(* Logix 5000 project; controller MV vendor 1 type 14 code 217 rev 31.11; software revision 31.00; part 45 of 53 *)
(* tags used below, declared in another part *)
   Always_Off : BOOL;
   CWD : CHECKWORD_FLAGS;
   Enable_TimeString : BOOL;
   MV22_TP_Capture_Volume_Timer : TIMER;
   MV_BM01_AV01 : PlantItem;   // BM01_AV01
   MV_BM01_AV01_CIP : BOOL;
   MV_BM01_AV01_MV21 : BOOL;
   MV_DAL01_AV01_MV21 : BOOL;
   MV_Enable_MV21_NewPressureControl : BOOL;
   MV_Enable_MV22_NewPressureControl : BOOL;
   MV_GasAvailable : BOOL;
   MV_MV21_AV01 : PlantItem;   // MV21_AV01
   MV_MV21_CIP : BOOL;
   MV_MV21_CO2 : BOOL;
   MV_MV21_CO2_ON_PreStorage : BOOL;
   MV_MV21_CO2_ON_Storage : BOOL;
   MV_MV21_ControlOpenVent : BOOL;
   MV_MV21_Filling_Pulse : BOOL;
   MV_MV21_Filling_PulseLevel : REAL;
   MV_MV21_LTX07_TrueLevel : REAL;
   MV_MV21_ProxiesOK : BOOL;
   MV_MV21_PTX01_AI : PlantItem;   // MV21_PTX01
   MV_MV21_TP_CaskDepressure : BOOL;
   MV_MV21_TP_CaskEmptying : BOOL;
   MV_MV21_TP_CaskFilling : BOOL;
   MV_MV21_TP_CaskPrePressure : BOOL;
   MV_MV21_TP_CaskReadyToFill : BOOL;
   MV_MV21_TP_CaskStorage : BOOL;
   MV_MV21_TP_CO2_Debounce_Timer : TIMER;
   MV_MV21_TP_CO2_Debounce_Timer_1 : TIMER;
   MV_MV21_TP_CO2_HSL_Pressure : REAL;
   MV_MV21_TP_CO2_HSL_Storage : REAL;
   MV_MV21_TP_CO2_HSL_Timer : TIMER;
   MV_MV21_TP_CO2_LSL_pressure_1 : REAL;
   MV_MV21_TP_CO2_LSL_storage : REAL;
   MV_MV21_TP_CO2_LSL_Timer : TIMER;
   MV_MV21_TP_Command : DINT;
   MV_MV21_TP_DAL_Chase_Cask : BOOL;
   MV_MV21_TP_DAL_Chase_KB : BOOL;
   MV_MV21_TP_DAL_Chase_Time : TIMER;
   MV_MV21_TP_Error_String : STRING;
   MV_MV21_TP_Faulted : BOOL;
   MV_MV21_TP_Fill_Pulse_OFF_Timer : TIMER;
   MV_MV21_TP_Fill_Pulse_ON_Timer : TIMER;
   MV_MV21_TP_Held : BOOL;
   MV_MV21_TP_Idle : BOOL;
   MV_MV21_TP_Initial_DAL_Chase_Cask : BOOL;
   MV_MV21_TP_Initial_DAL_Chase_KB : BOOL;
   MV_MV21_TP_KBEmptying : BOOL;
   MV_MV21_TP_KBFilling : BOOL;
   MV_MV21_TP_KBFillingBuildPressure : BOOL;
   MV_MV21_TP_KBPreEmptyPressure : BOOL;
   MV_MV21_TP_KBPrePressurise : BOOL;
   MV_MV21_TP_KBStorage : BOOL;
   MV_MV21_TP_LowerLimit : REAL;
   MV_MV21_TP_NotIdle : BOOL;
   MV_MV21_TP_Prompt : DINT;
   MV_MV21_TP_Pulse : BOOL;
   MV_MV21_TP_ReadyToFillKB : BOOL;
   MV_MV21_TP_ReadyToFillKB_M : BOOL;
   MV_MV21_TP_Running : BOOL;
   MV_MV21_TP_Setpoint : REAL;
   MV_MV21_TP_Status : DINT;   // 0 = Idle, 1 = Running, 2 = Held, 3 = Faulted
   MV_MV21_TP_Step : DINT;
   MV_MV21_TP_Steptime : DINT;
   MV_MV21_TP_Steptime_String : STRING;
   MV_MV21_TP_SteptimeRunning : DINT;
   MV_MV21_TP_TimeLeft : DINT;
   MV_MV21_TP_TimeLeft_msec : DINT;
   MV_MV21_TP_TimeLeftStr : STRING;
   MV_MV21_TP_UpperLimit : REAL;
   MV_MV21_TP_Vent : BOOL;
   MV_MV21_TPLastStep : DINT;
   MV_MV22_CO2_ON_PreStorage : BOOL;
   MV_MV22_CO2_ON_Storage : BOOL;
   MV_MV22_Filling_PulseLevel : DINT;
   MV_MV22_LTX07_TrueLevel : REAL;
   MV_MV22_ProxiesOK : BOOL;
   MV_MV22_PTX01_AI : PlantItem;   // MV22_PTX01
   MV_MV22_TP_CaskPurgeFromTop : BOOL;
   MV_MV22_TP_Command : DINT;
   MV_MV22_TP_DAL_Chase_KB : BOOL;
   MV_MV22_TP_Dirty : BOOL;
   MV_MV22_TP_Emptying_Level_Setpoint : REAL;
   MV_MV22_TP_Idle : BOOL;
   MV_MV22_TP_Initial_DAL_Chase_KB : BOOL;
   MV_MV22_TP_KBDepressure : BOOL;
   MV_MV22_TP_KBEmptying : BOOL;
   MV_MV22_TP_KBFilling : BOOL;
   MV_MV22_TP_KBFilling_M : BOOL;
   MV_MV22_TP_KBPreEmptyPressure : BOOL;
   MV_MV22_TP_KBPrePressurise : BOOL;
   MV_MV22_TP_KBPurgeFromTop : BOOL;
   MV_MV22_TP_KBPurgeTimer : TIMER;
   MV_MV22_TP_KBStorage : BOOL;
   MV_MV22_TP_ONS : BOOL;
   MV_MV22_TP_Prompt : DINT;
   MV_MV22_TP_ReadyToFillKB : BOOL;
   MV_MV22_TP_ReadyToFillKB_M : BOOL;
   MV_MV22_TP_Running : BOOL;
   MV_MV22_TP_Setpoint : REAL;
   MV_MV22_TP_Status : DINT;   // 0 = Idle, 1 = Running, 2 = Held, 3 = Faulted
   MV_MV22_TP_Step : DINT;
   MV_MV22_TP_Steptime : DINT;
   MV_MV22_TP_UpperLimit : REAL;
   MV_MV22_Transfer_StartLevel : REAL;
   MV_MV22_Transferred_Level : REAL;
   MV_N138 : INT[50];   // MV 22, CURRENT FV DATA
   MV_TP_CaskFillingPressure : REAL;
   MV_TP_CaskPrefillPressure : REAL;
   MV_TP_CaskStoragePressure : REAL;
   MV_TP_CaskStoragePressureDelay_Secs : DINT;
   MV_TP_Deadband : REAL;
   MV_TP_Emptying_Volume_Setpoint : REAL;
   MV_TP_HighLevelDeadband : REAL;
   MV_TP_KBEmptyingPressure : REAL;
   MV_TP_KBFillingPressure : REAL;
   MV_TP_KBPrefillPressure : REAL;
   MV_TP_KBStoragePressure : REAL;
   MV_TP_KBStoragePressureLevel : REAL;
   MV_TP_LowLevelDeadbandThreshold : REAL;
   MV_TP_NoCIPDelay : DINT;
   One_Second_1_scan : BOOL;
(* MV_Common, continued *)

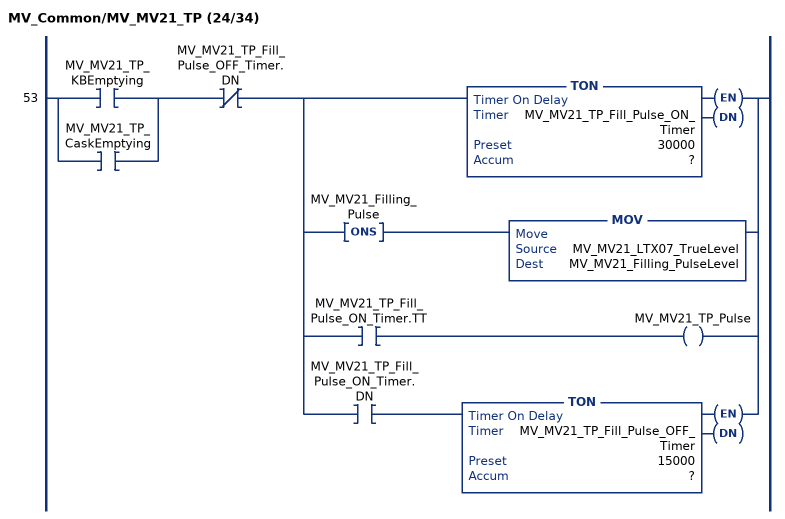
   53: [XIC(MV_MV21_TP_KBEmptying) ,XIC(MV_MV21_TP_CaskEmptying) ]XIO(MV_MV21_TP_Fill_Pulse_OFF_Timer.DN)[TON(MV_MV21_TP_Fill_Pulse_ON_Timer,?,?) ,ONS(MV_MV21_Filling_Pulse) MOV(MV_MV21_LTX07_TrueLevel,MV_MV21_Filling_PulseLevel) ,XIC(MV_MV21_TP_Fill_Pulse_ON_Timer.TT) OTE(MV_MV21_TP_Pulse) ,XIC(MV_MV21_TP_Fill_Pulse_ON_Timer.DN) TON(MV_MV21_TP_Fill_Pulse_OFF_Timer,?,?) ];
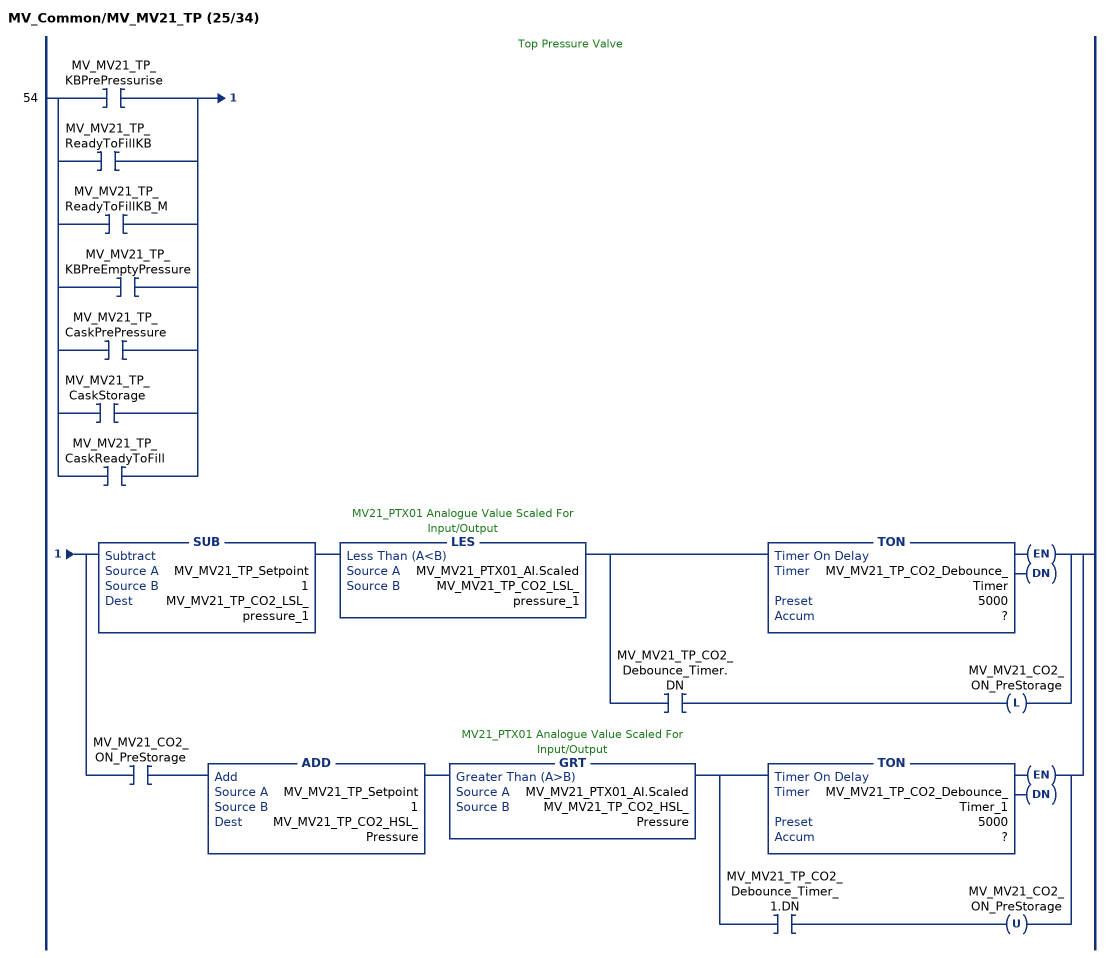
   // Top Pressure Valve
   54: [XIC(MV_MV21_TP_KBPrePressurise) ,XIC(MV_MV21_TP_ReadyToFillKB) ,XIC(MV_MV21_TP_ReadyToFillKB_M) ,XIC(MV_MV21_TP_KBPreEmptyPressure) ,XIC(MV_MV21_TP_CaskPrePressure) ,XIC(MV_MV21_TP_CaskStorage) ,XIC(MV_MV21_TP_CaskReadyToFill) ][SUB(MV_MV21_TP_Setpoint,1,MV_MV21_TP_CO2_LSL_pressure_1) LES(MV_MV21_PTX01_AI.Scaled,MV_MV21_TP_CO2_LSL_pressure_1) [TON(MV_MV21_TP_CO2_Debounce_Timer,?,?) ,XIC(MV_MV21_TP_CO2_Debounce_Timer.DN) OTL(MV_MV21_CO2_ON_PreStorage) ] ,XIC(MV_MV21_CO2_ON_PreStorage) ADD(MV_MV21_TP_Setpoint,1,MV_MV21_TP_CO2_HSL_Pressure) GRT(MV_MV21_PTX01_AI.Scaled,MV_MV21_TP_CO2_HSL_Pressure) [TON(MV_MV21_TP_CO2_Debounce_Timer_1,?,?) ,XIC(MV_MV21_TP_CO2_Debounce_Timer_1.DN) OTU(MV_MV21_CO2_ON_PreStorage) ] ];
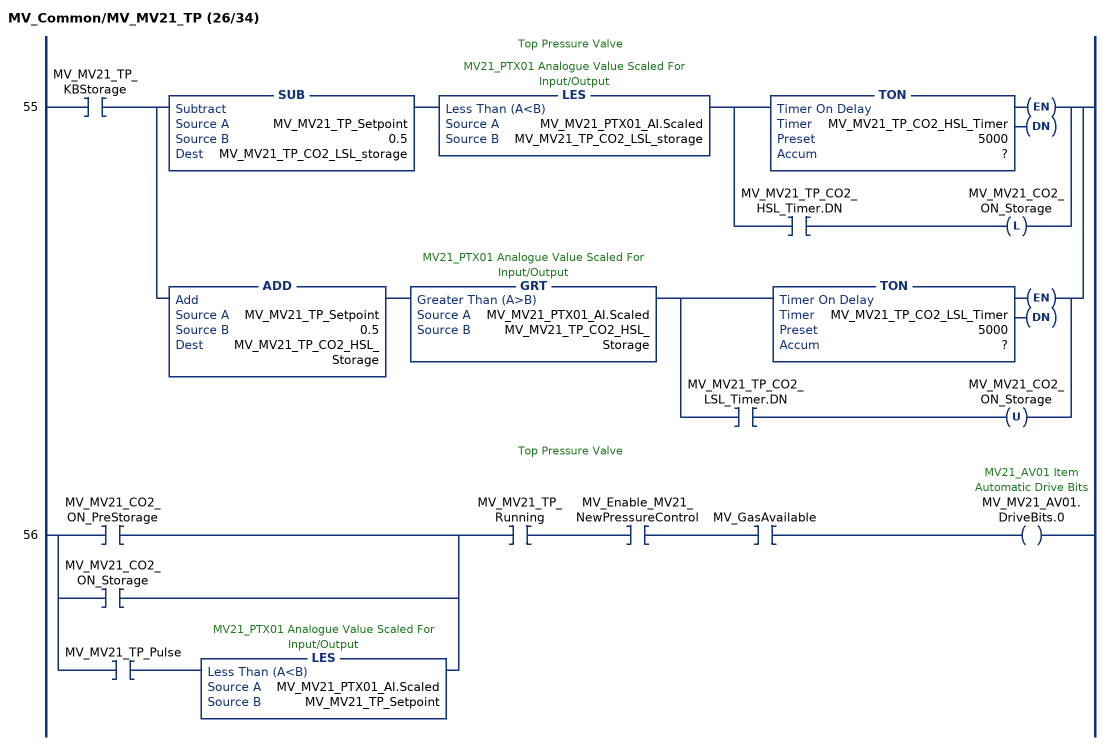
   // Top Pressure Valve
   55: XIC(MV_MV21_TP_KBStorage)[SUB(MV_MV21_TP_Setpoint,0.5,MV_MV21_TP_CO2_LSL_storage) LES(MV_MV21_PTX01_AI.Scaled,MV_MV21_TP_CO2_LSL_storage) [TON(MV_MV21_TP_CO2_HSL_Timer,?,?) ,XIC(MV_MV21_TP_CO2_HSL_Timer.DN) OTL(MV_MV21_CO2_ON_Storage) ] ,ADD(MV_MV21_TP_Setpoint,0.5,MV_MV21_TP_CO2_HSL_Storage) GRT(MV_MV21_PTX01_AI.Scaled,MV_MV21_TP_CO2_HSL_Storage) [TON(MV_MV21_TP_CO2_LSL_Timer,?,?) ,XIC(MV_MV21_TP_CO2_LSL_Timer.DN) OTU(MV_MV21_CO2_ON_Storage) ] ];
   // Top Pressure Valve
   56: [XIC(MV_MV21_CO2_ON_PreStorage) ,XIC(MV_MV21_CO2_ON_Storage) ,XIC(MV_MV21_TP_Pulse) LES(MV_MV21_PTX01_AI.Scaled,MV_MV21_TP_Setpoint) ]XIC(MV_MV21_TP_Running)XIC(MV_Enable_MV21_NewPressureControl)XIC(MV_GasAvailable)OTE(MV_MV21_AV01.DriveBits.0);
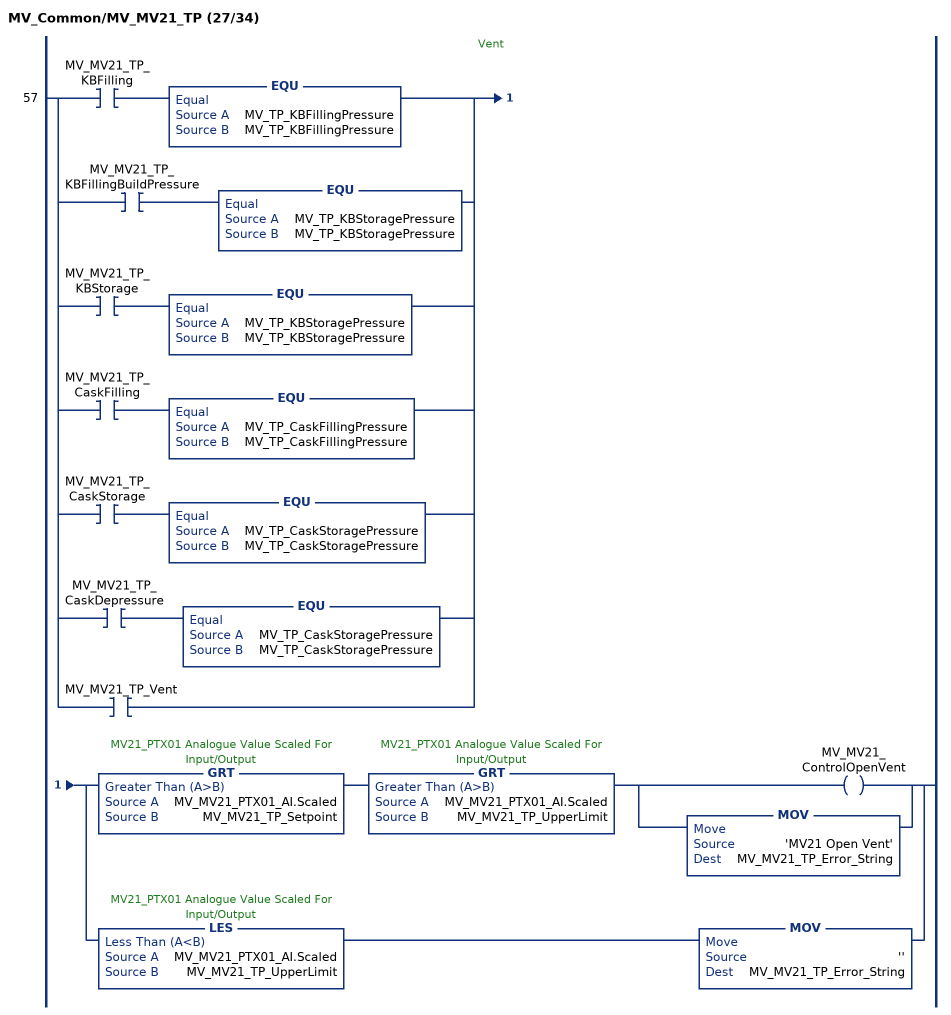
   // Vent
   57: [XIC(MV_MV21_TP_KBFilling) EQU(MV_TP_KBFillingPressure,MV_TP_KBFillingPressure) ,XIC(MV_MV21_TP_KBFillingBuildPressure) EQU(MV_TP_KBStoragePressure,MV_TP_KBStoragePressure) ,XIC(MV_MV21_TP_KBStorage) EQU(MV_TP_KBStoragePressure,MV_TP_KBStoragePressure) ,XIC(MV_MV21_TP_CaskFilling) EQU(MV_TP_CaskFillingPressure,MV_TP_CaskFillingPressure) ,XIC(MV_MV21_TP_CaskStorage) EQU(MV_TP_CaskStoragePressure,MV_TP_CaskStoragePressure) ,XIC(MV_MV21_TP_CaskDepressure) EQU(MV_TP_CaskStoragePressure,MV_TP_CaskStoragePressure) ,XIC(MV_MV21_TP_Vent) ][GRT(MV_MV21_PTX01_AI.Scaled,MV_MV21_TP_Setpoint) GRT(MV_MV21_PTX01_AI.Scaled,MV_MV21_TP_UpperLimit) [OTE(MV_MV21_ControlOpenVent) ,MOV('MV21 Open Vent',MV_MV21_TP_Error_String) ] ,LES(MV_MV21_PTX01_AI.Scaled,MV_MV21_TP_UpperLimit) MOV('',MV_MV21_TP_Error_String) ];
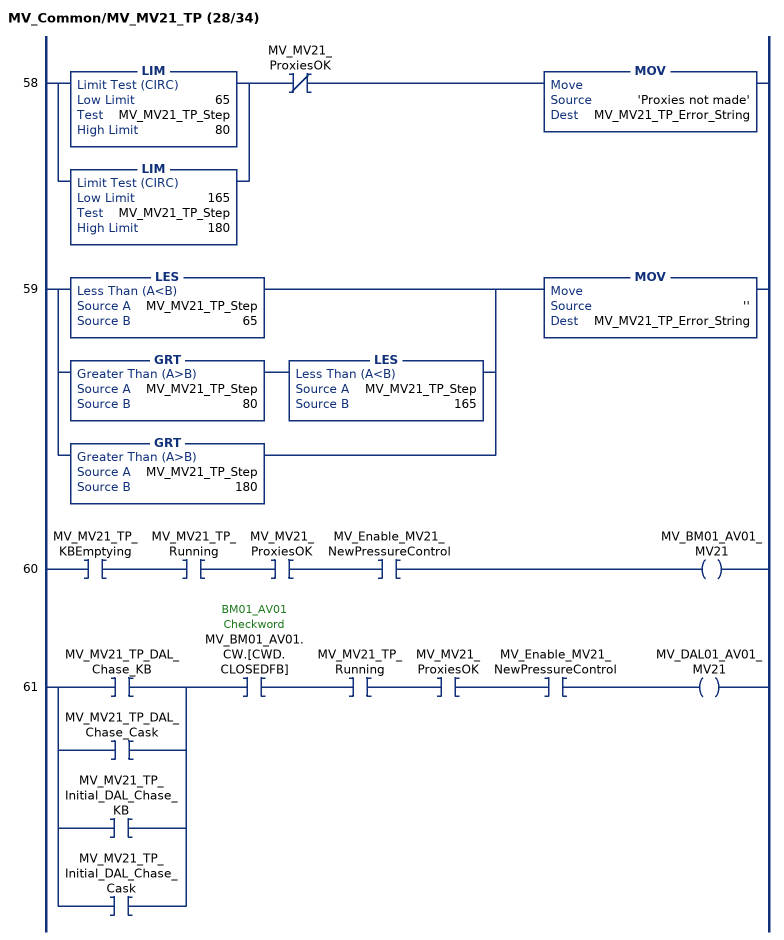
   58: [LIM(65,MV_MV21_TP_Step,80) ,LIM(165,MV_MV21_TP_Step,180) ]XIO(MV_MV21_ProxiesOK)MOV('Proxies not made',MV_MV21_TP_Error_String);
   59: [LES(MV_MV21_TP_Step,65) ,GRT(MV_MV21_TP_Step,80) LES(MV_MV21_TP_Step,165) ,GRT(MV_MV21_TP_Step,180) ]MOV('',MV_MV21_TP_Error_String);
   60: XIC(MV_MV21_TP_KBEmptying)XIC(MV_MV21_TP_Running)XIC(MV_MV21_ProxiesOK)XIC(MV_Enable_MV21_NewPressureControl)OTE(MV_BM01_AV01_MV21);
   61: [XIC(MV_MV21_TP_DAL_Chase_KB) ,XIC(MV_MV21_TP_DAL_Chase_Cask) ,XIC(MV_MV21_TP_Initial_DAL_Chase_KB) ,XIC(MV_MV21_TP_Initial_DAL_Chase_Cask) ]XIC(MV_BM01_AV01.CW.[CWD.CLOSEDFB])XIC(MV_MV21_TP_Running)XIC(MV_MV21_ProxiesOK)XIC(MV_Enable_MV21_NewPressureControl)OTE(MV_DAL01_AV01_MV21);
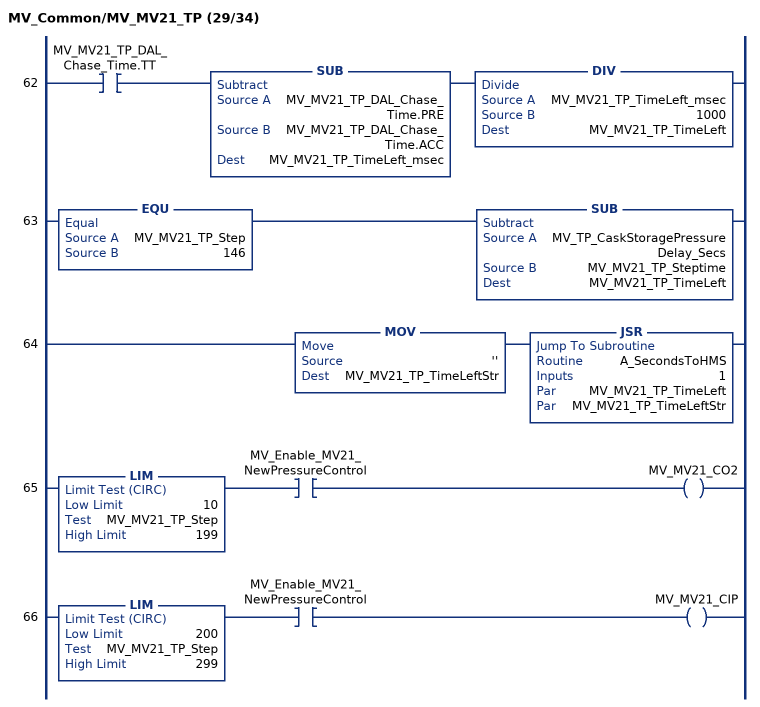
   62: XIC(MV_MV21_TP_DAL_Chase_Time.TT)SUB(MV_MV21_TP_DAL_Chase_Time.PRE,MV_MV21_TP_DAL_Chase_Time.ACC,MV_MV21_TP_TimeLeft_msec)DIV(MV_MV21_TP_TimeLeft_msec,1000,MV_MV21_TP_TimeLeft);
   63: EQU(MV_MV21_TP_Step,146)SUB(MV_TP_CaskStoragePressureDelay_Secs,MV_MV21_TP_Steptime,MV_MV21_TP_TimeLeft);
   64: MOV('',MV_MV21_TP_TimeLeftStr)JSR(A_SecondsToHMS,1,MV_MV21_TP_TimeLeft,MV_MV21_TP_TimeLeftStr);
   65: LIM(10,MV_MV21_TP_Step,199)XIC(MV_Enable_MV21_NewPressureControl)OTE(MV_MV21_CO2);
   66: LIM(200,MV_MV21_TP_Step,299)XIC(MV_Enable_MV21_NewPressureControl)OTE(MV_MV21_CIP);
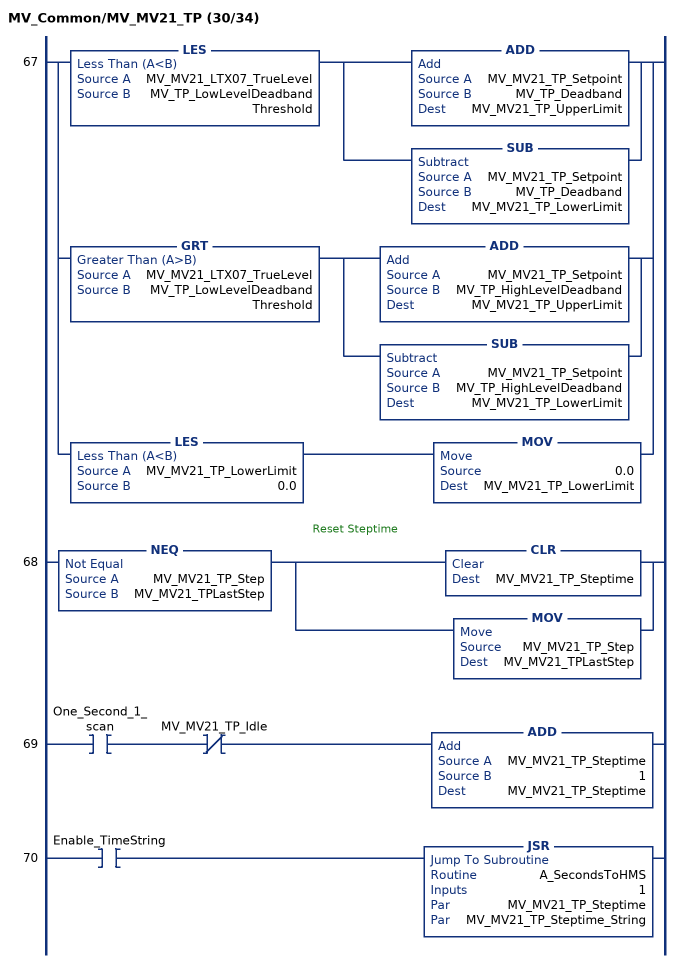
   67: [LES(MV_MV21_LTX07_TrueLevel,MV_TP_LowLevelDeadbandThreshold) [ADD(MV_MV21_TP_Setpoint,MV_TP_Deadband,MV_MV21_TP_UpperLimit) ,SUB(MV_MV21_TP_Setpoint,MV_TP_Deadband,MV_MV21_TP_LowerLimit) ] ,GRT(MV_MV21_LTX07_TrueLevel,MV_TP_LowLevelDeadbandThreshold) [ADD(MV_MV21_TP_Setpoint,MV_TP_HighLevelDeadband,MV_MV21_TP_UpperLimit) ,SUB(MV_MV21_TP_Setpoint,MV_TP_HighLevelDeadband,MV_MV21_TP_LowerLimit) ] ,LES(MV_MV21_TP_LowerLimit,0.0) MOV(0.0,MV_MV21_TP_LowerLimit) ];
   // Reset Steptime
   68: NEQ(MV_MV21_TP_Step,MV_MV21_TPLastStep)[CLR(MV_MV21_TP_Steptime) ,MOV(MV_MV21_TP_Step,MV_MV21_TPLastStep) ];
   69: XIC(One_Second_1_scan)XIO(MV_MV21_TP_Idle)ADD(MV_MV21_TP_Steptime,1,MV_MV21_TP_Steptime);
   70: XIC(Enable_TimeString)JSR(A_SecondsToHMS,1,MV_MV21_TP_Steptime,MV_MV21_TP_Steptime_String);
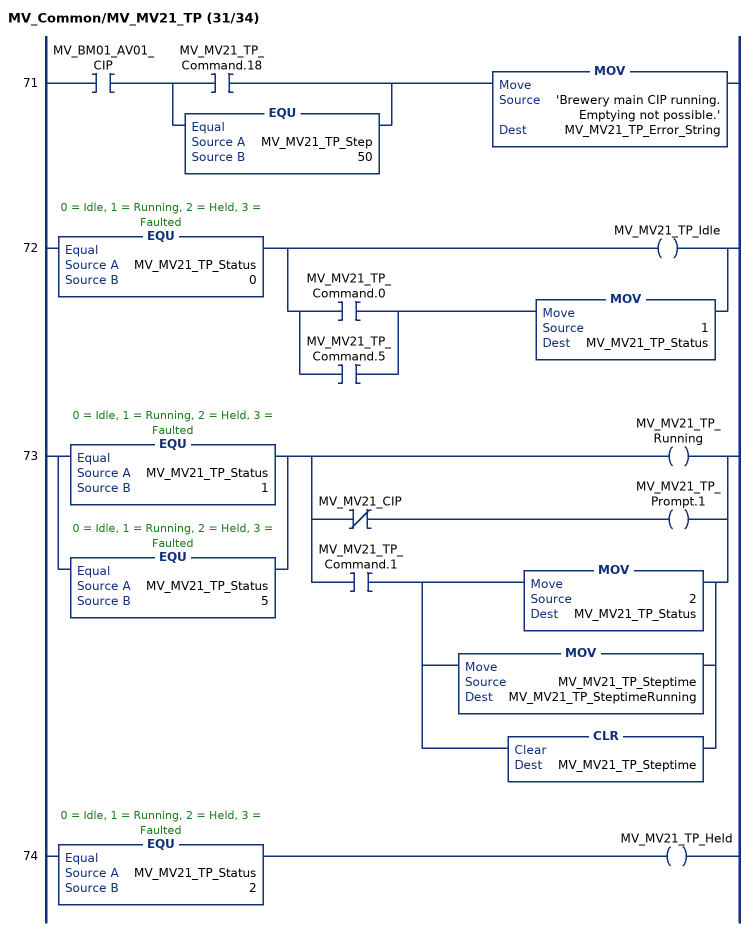
   71: XIC(MV_BM01_AV01_CIP)[XIC(MV_MV21_TP_Command.18) ,EQU(MV_MV21_TP_Step,50) ]MOV('Brewery main CIP running. Emptying not possible.',MV_MV21_TP_Error_String);
   72: EQU(MV_MV21_TP_Status,0)[OTE(MV_MV21_TP_Idle) ,[XIC(MV_MV21_TP_Command.0) ,XIC(MV_MV21_TP_Command.5) ] MOV(1,MV_MV21_TP_Status) ];
   73: [EQU(MV_MV21_TP_Status,1) ,EQU(MV_MV21_TP_Status,5) ][OTE(MV_MV21_TP_Running) ,XIO(MV_MV21_CIP) OTE(MV_MV21_TP_Prompt.1) ,XIC(MV_MV21_TP_Command.1) [MOV(2,MV_MV21_TP_Status) ,MOV(MV_MV21_TP_Steptime,MV_MV21_TP_SteptimeRunning) ,CLR(MV_MV21_TP_Steptime) ] ];
   74: EQU(MV_MV21_TP_Status,2)OTE(MV_MV21_TP_Held);
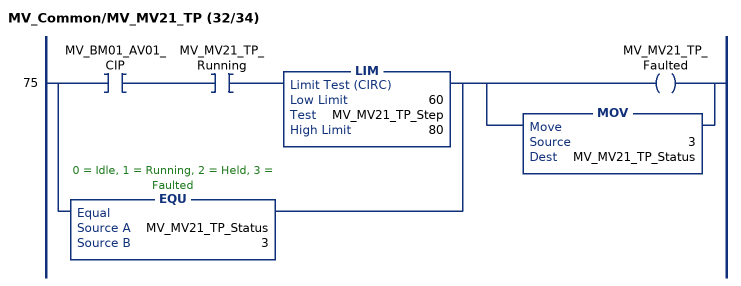
   75: [XIC(MV_BM01_AV01_CIP) XIC(MV_MV21_TP_Running) LIM(60,MV_MV21_TP_Step,80) ,EQU(MV_MV21_TP_Status,3) ][OTE(MV_MV21_TP_Faulted) ,MOV(3,MV_MV21_TP_Status) ];
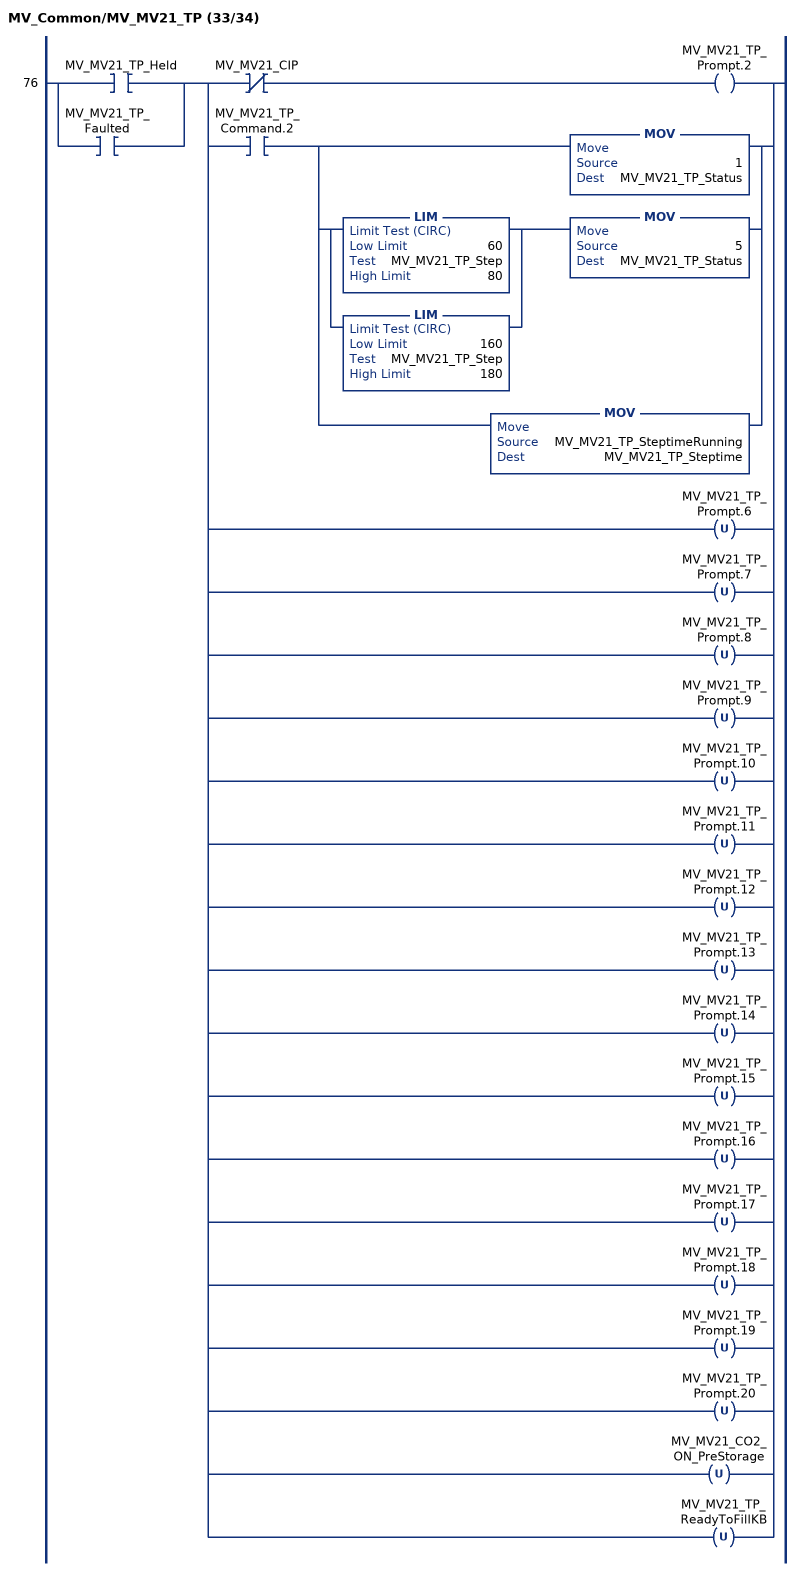
   76: [XIC(MV_MV21_TP_Held) ,XIC(MV_MV21_TP_Faulted) ][XIO(MV_MV21_CIP) OTE(MV_MV21_TP_Prompt.2) ,XIC(MV_MV21_TP_Command.2) [MOV(1,MV_MV21_TP_Status) ,[LIM(60,MV_MV21_TP_Step,80) ,LIM(160,MV_MV21_TP_Step,180) ] MOV(5,MV_MV21_TP_Status) ,MOV(MV_MV21_TP_SteptimeRunning,MV_MV21_TP_Steptime) ] ,OTU(MV_MV21_TP_Prompt.6) ,OTU(MV_MV21_TP_Prompt.7) ,OTU(MV_MV21_TP_Prompt.8) ,OTU(MV_MV21_TP_Prompt.9) ,OTU(MV_MV21_TP_Prompt.10) ,OTU(MV_MV21_TP_Prompt.11) ,OTU(MV_MV21_TP_Prompt.12) ,OTU(MV_MV21_TP_Prompt.13) ,OTU(MV_MV21_TP_Prompt.14) ,OTU(MV_MV21_TP_Prompt.15) ,OTU(MV_MV21_TP_Prompt.16) ,OTU(MV_MV21_TP_Prompt.17) ,OTU(MV_MV21_TP_Prompt.18) ,OTU(MV_MV21_TP_Prompt.19) ,OTU(MV_MV21_TP_Prompt.20) ,OTU(MV_MV21_CO2_ON_PreStorage) ,OTU(MV_MV21_TP_ReadyToFillKB) ];